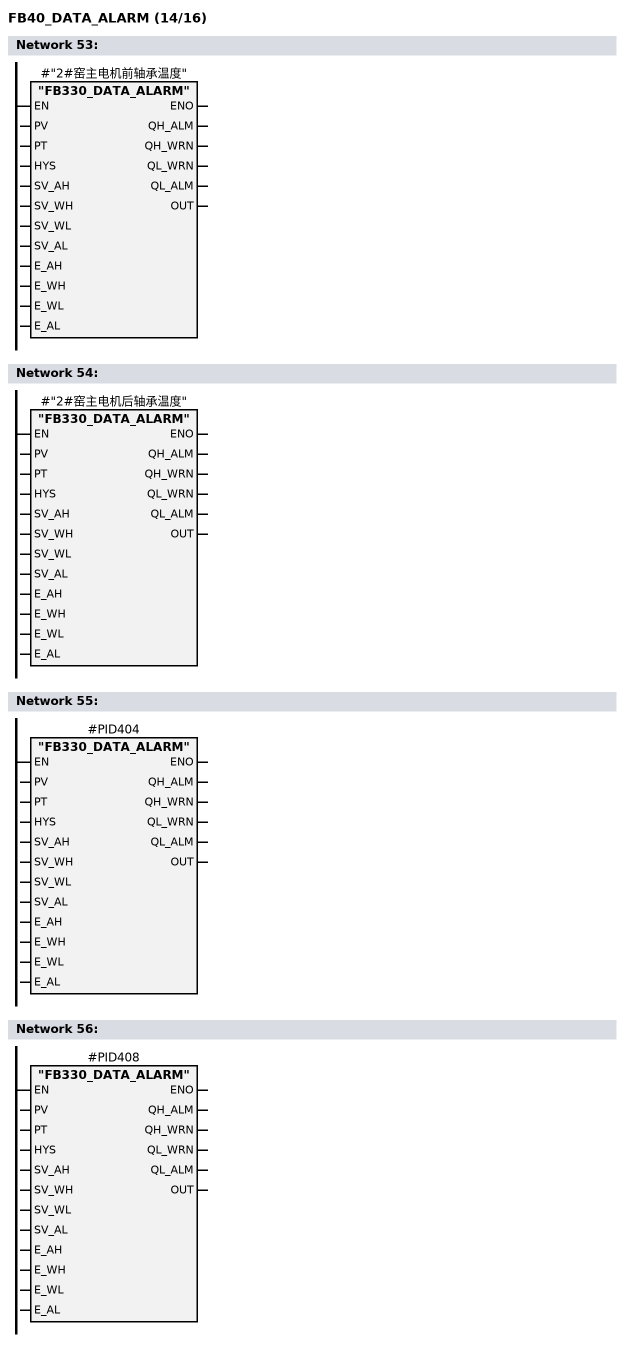
   RUNG wire#powerrail
      #"2#窑主电机前轴承温度"(PV :=, PT :=, HYS :=, SV_AH :=, SV_WH :=, SV_WL :=, SV_AL :=, E_AH :=, E_WH :=, E_WL :=, E_AL :=, QH_ALM =>, QH_WRN =>, QL_WRN =>, QL_ALM =>, OUT =>)
   END_RUNG
   // the same network as SCL:
   #"2#窑主电机前轴承温度"();   // "FB330_DATA_ALARM"
END_REGION

REGION Network 54
   RUNG wire#powerrail
      #"2#窑主电机后轴承温度"(PV :=, PT :=, HYS :=, SV_AH :=, SV_WH :=, SV_WL :=, SV_AL :=, E_AH :=, E_WH :=, E_WL :=, E_AL :=, QH_ALM =>, QH_WRN =>, QL_WRN =>, QL_ALM =>, OUT =>)
   END_RUNG
   // the same network as SCL:
   #"2#窑主电机后轴承温度"();   // "FB330_DATA_ALARM"
END_REGION

REGION Network 55
   RUNG wire#powerrail
      #PID404(PV :=, PT :=, HYS :=, SV_AH :=, SV_WH :=, SV_WL :=, SV_AL :=, E_AH :=, E_WH :=, E_WL :=, E_AL :=, QH_ALM =>, QH_WRN =>, QL_WRN =>, QL_ALM =>, OUT =>)
   END_RUNG
   // the same network as SCL:
   #PID404();   // "FB330_DATA_ALARM"
END_REGION

REGION Network 56
   RUNG wire#powerrail
      #PID408(PV :=, PT :=, HYS :=, SV_AH :=, SV_WH :=, SV_WL :=, SV_AL :=, E_AH :=, E_WH :=, E_WL :=, E_AL :=, QH_ALM =>, QH_WRN =>, QL_WRN =>, QL_ALM =>, OUT =>)
   END_RUNG
   // the same network as SCL:
   #PID408();   // "FB330_DATA_ALARM"
END_REGION

REGION Network 57
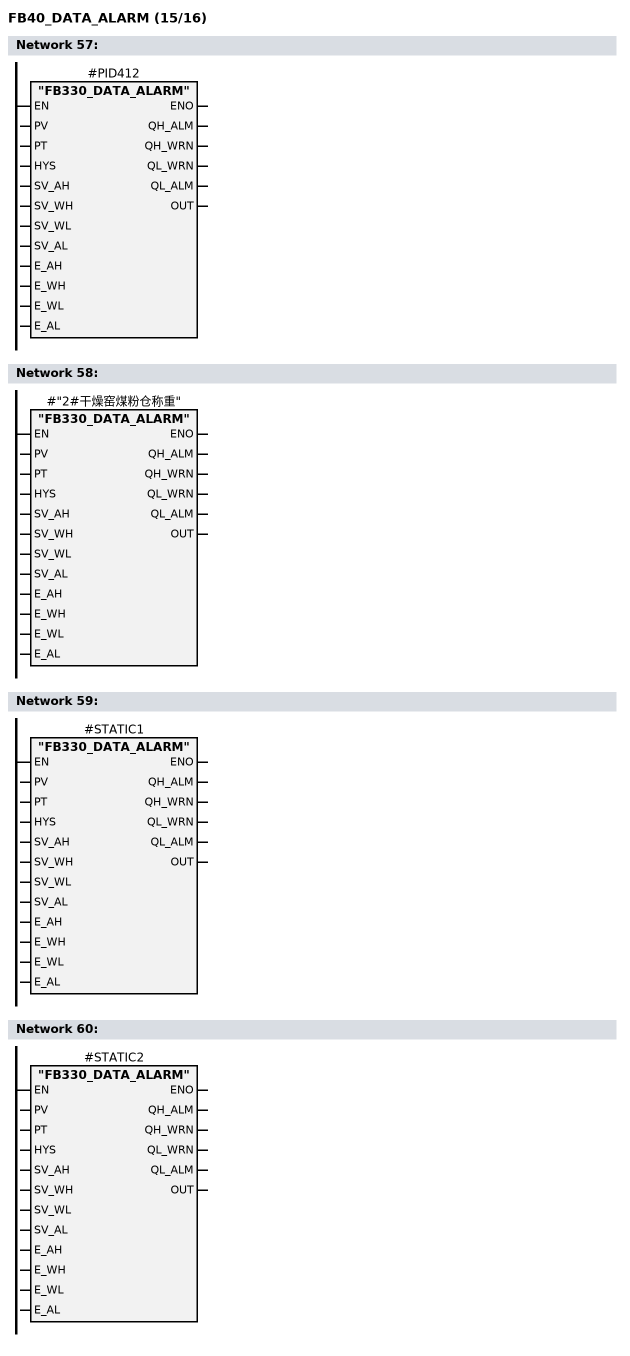
   RUNG wire#powerrail
      #PID412(PV :=, PT :=, HYS :=, SV_AH :=, SV_WH :=, SV_WL :=, SV_AL :=, E_AH :=, E_WH :=, E_WL :=, E_AL :=, QH_ALM =>, QH_WRN =>, QL_WRN =>, QL_ALM =>, OUT =>)
   END_RUNG
   // the same network as SCL:
   #PID412();   // "FB330_DATA_ALARM"
END_REGION

REGION Network 58
   RUNG wire#powerrail
      #"2#干燥窑煤粉仓称重"(PV :=, PT :=, HYS :=, SV_AH :=, SV_WH :=, SV_WL :=, SV_AL :=, E_AH :=, E_WH :=, E_WL :=, E_AL :=, QH_ALM =>, QH_WRN =>, QL_WRN =>, QL_ALM =>, OUT =>)
   END_RUNG
   // the same network as SCL:
   #"2#干燥窑煤粉仓称重"();   // "FB330_DATA_ALARM"
END_REGION

REGION Network 59
   RUNG wire#powerrail
      #STATIC1(PV :=, PT :=, HYS :=, SV_AH :=, SV_WH :=, SV_WL :=, SV_AL :=, E_AH :=, E_WH :=, E_WL :=, E_AL :=, QH_ALM =>, QH_WRN =>, QL_WRN =>, QL_ALM =>, OUT =>)
   END_RUNG
   // the same network as SCL:
   #STATIC1();   // "FB330_DATA_ALARM"
END_REGION

REGION Network 60
   RUNG wire#powerrail
      #STATIC2(PV :=, PT :=, HYS :=, SV_AH :=, SV_WH :=, SV_WL :=, SV_AL :=, E_AH :=, E_WH :=, E_WL :=, E_AL :=, QH_ALM =>, QH_WRN =>, QL_WRN =>, QL_ALM =>, OUT =>)
   END_RUNG
   // the same network as SCL:
   #STATIC2();   // "FB330_DATA_ALARM"
END_REGION

REGION Network 61
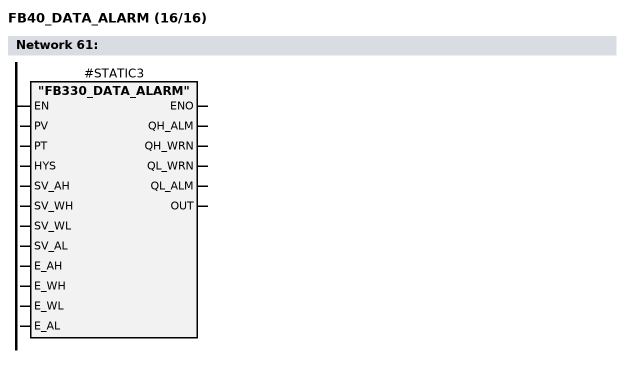
   RUNG wire#powerrail
      #STATIC3(PV :=, PT :=, HYS :=, SV_AH :=, SV_WH :=, SV_WL :=, SV_AL :=, E_AH :=, E_WH :=, E_WL :=, E_AL :=, QH_ALM =>, QH_WRN =>, QL_WRN =>, QL_ALM =>, OUT =>)
   END_RUNG
   // the same network as SCL:
   #STATIC3();   // "FB330_DATA_ALARM"
END_REGION
END_FUNCTION_BLOCK

FUNCTION_BLOCK "FB330_DATA_ALARM"   // FB330, LAD
{ S7_Optimized_Access := 'FALSE' }
VERSION : 0.1
// REAL的报警块
   VAR_INPUT
      PV : Real;   // 过程值
      PT : Real := 1.0;   // 系数
      HYS : Real;   // 回差值
      SV_AH : Real;   // 高报警设定值
      SV_WH : Real;   // 高警告设定值
      SV_WL : Real;   // 低警告设定值
      SV_AL : Real;   // 低报警设定值
      E_AH : Bool;   // 高报警使能
      E_WH : Bool;   // 高警告使能
      E_WL : Bool;   // 低警告使能
      E_AL : Bool;   // 低报警使能
   END_VAR
   VAR_OUTPUT
      QH_ALM : Bool;   // 高报警输出
      QH_WRN : Bool;   // 高警告输出
      QL_WRN : Bool;   // 低警告输出
      QL_ALM : Bool;   // 低报警输出
      OUT : Real;   // 输出
   END_VAR
   VAR
      SR1 : Bool;
      SR2 : Bool;
      SR3 : Bool;
      SR4 : Bool;
   END_VAR
   VAR_TEMP
      TEMP_AH : Real;
      TEMP_WH : Real;
      TEMP_AL : Real;
      TEMP_WL : Real;
      TEMP_OUT : Real;
   END_VAR
BEGIN

REGION Network 1
   // 系数转换
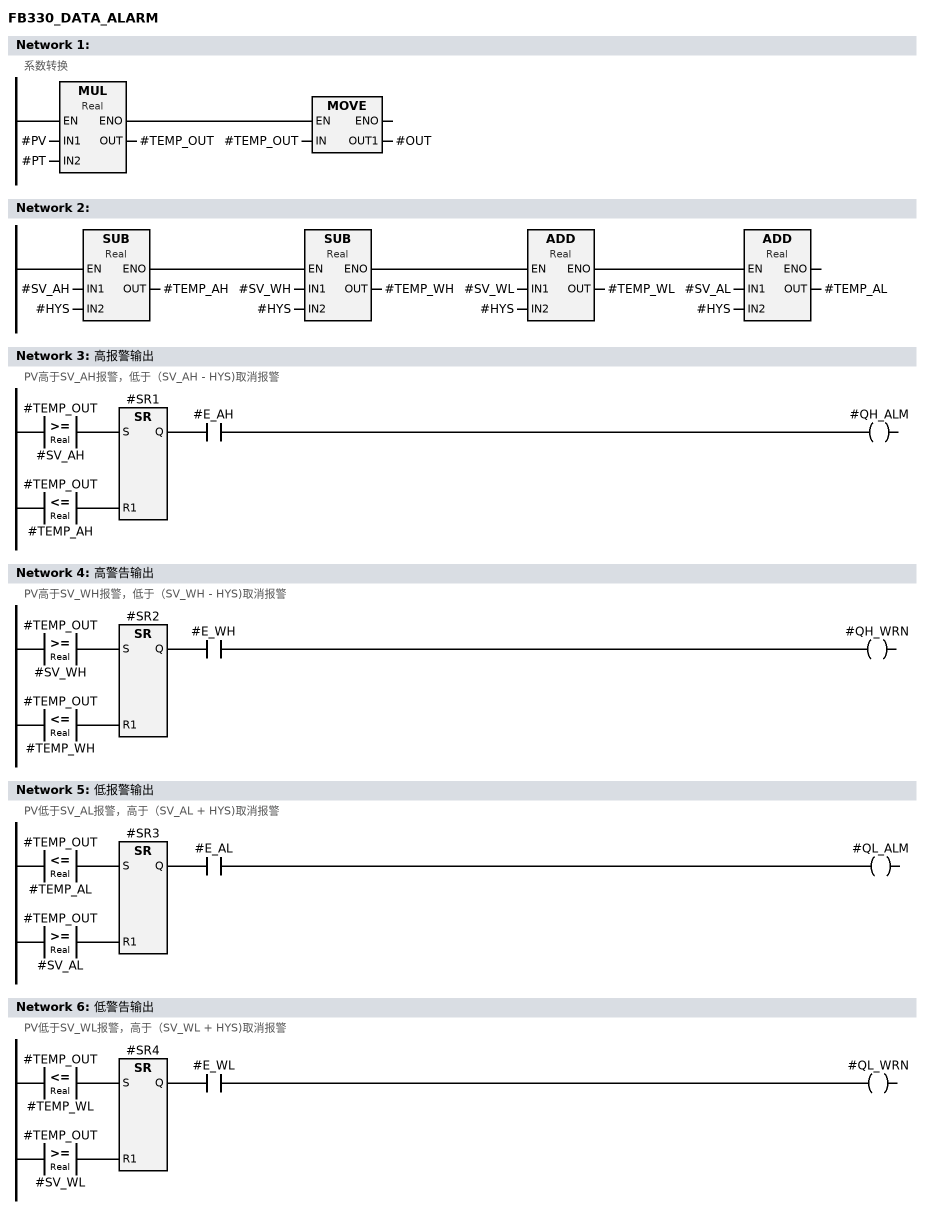
   RUNG wire#powerrail
      { S7_Templates := "SrcType := Real"; S7_GenerateENO := "TRUE" } Mul(in1 := #PV, in2 := #PT, out => #TEMP_OUT)
      { S7_GenerateENO := "TRUE" } Move(in := #TEMP_OUT, out1 => #OUT)
   END_RUNG
   // the same network as SCL:
   // ENO of a box is taken as its EN; it also drops when the box reports an error
   #TEMP_OUT := #PV * #PT;
   #OUT := #TEMP_OUT;
END_REGION

REGION Network 2
   RUNG wire#powerrail
      { S7_Templates := "SrcType := Real"; S7_GenerateENO := "TRUE" } Sub(in1 := #SV_AH, in2 := #HYS, out => #TEMP_AH)
      { S7_Templates := "SrcType := Real"; S7_GenerateENO := "TRUE" } Sub(in1 := #SV_WH, in2 := #HYS, out => #TEMP_WH)
      { S7_Templates := "SrcType := Real"; S7_GenerateENO := "TRUE" } Add(in1 := #SV_WL, in2 := #HYS, out => #TEMP_WL)
      { S7_Templates := "SrcType := Real"; S7_GenerateENO := "TRUE" } Add(in1 := #SV_AL, in2 := #HYS, out => #TEMP_AL)
   END_RUNG
   // the same network as SCL:
   // ENO of a box is taken as its EN; it also drops when the box reports an error
   #TEMP_AH := #SV_AH - #HYS;
   #TEMP_WH := #SV_WH - #HYS;
   #TEMP_WL := #SV_WL + #HYS;
   #TEMP_AL := #SV_AL + #HYS;
END_REGION

REGION Network 3: 高报警输出
   // PV高于SV_AH报警，低于（SV_AH - HYS)取消报警
   RUNG wire#powerrail
      { S7_Templates := "SrcType := Real" } GE_Contact(in1 := #TEMP_OUT, in2 := #SV_AH)
      S_SR(operand := #SR1, r1 := wire#w1)
      Contact( #E_AH )
      Coil( #QH_ALM )
   END_RUNG
   RUNG wire#powerrail
      { S7_Templates := "SrcType := Real" } LE_Contact(in1 := #TEMP_OUT, in2 := #TEMP_AH)
   END_RUNG wire#w1
   // the same network as SCL:
   IF #TEMP_OUT >= #SV_AH THEN
       #SR1 := TRUE;   // SR flip-flop
   END_IF;
   IF #TEMP_OUT <= #TEMP_AH THEN #SR1 := FALSE; END_IF;
   #QH_ALM := #SR1 AND #E_AH;
END_REGION

REGION Network 4: 高警告输出
   // PV高于SV_WH报警，低于（SV_WH - HYS)取消报警
   RUNG wire#powerrail
      { S7_Templates := "SrcType := Real" } GE_Contact(in1 := #TEMP_OUT, in2 := #SV_WH)
      S_SR(operand := #SR2, r1 := wire#w1)
      Contact( #E_WH )
      Coil( #QH_WRN )
   END_RUNG
   RUNG wire#powerrail
      { S7_Templates := "SrcType := Real" } LE_Contact(in1 := #TEMP_OUT, in2 := #TEMP_WH)
   END_RUNG wire#w1
   // the same network as SCL:
   IF #TEMP_OUT >= #SV_WH THEN
       #SR2 := TRUE;   // SR flip-flop
   END_IF;
   IF #TEMP_OUT <= #TEMP_WH THEN #SR2 := FALSE; END_IF;
   #QH_WRN := #SR2 AND #E_WH;
END_REGION

REGION Network 5: 低报警输出
   // PV低于SV_AL报警，高于（SV_AL + HYS)取消报警
   RUNG wire#powerrail
      { S7_Templates := "SrcType := Real" } LE_Contact(in1 := #TEMP_OUT, in2 := #TEMP_AL)
      S_SR(operand := #SR3, r1 := wire#w1)
      Contact( #E_AL )
      Coil( #QL_ALM )
   END_RUNG
   RUNG wire#powerrail
      { S7_Templates := "SrcType := Real" } GE_Contact(in1 := #TEMP_OUT, in2 := #SV_AL)
   END_RUNG wire#w1
   // the same network as SCL:
   IF #TEMP_OUT <= #TEMP_AL THEN
       #SR3 := TRUE;   // SR flip-flop
   END_IF;
   IF #TEMP_OUT >= #SV_AL THEN #SR3 := FALSE; END_IF;
   #QL_ALM := #SR3 AND #E_AL;
END_REGION

REGION Network 6: 低警告输出
   // PV低于SV_WL报警，高于（SV_WL + HYS)取消报警
   RUNG wire#powerrail
      { S7_Templates := "SrcType := Real" } LE_Contact(in1 := #TEMP_OUT, in2 := #TEMP_WL)
      S_SR(operand := #SR4, r1 := wire#w1)
      Contact( #E_WL )
      Coil( #QL_WRN )
   END_RUNG
   RUNG wire#powerrail
      { S7_Templates := "SrcType := Real" } GE_Contact(in1 := #TEMP_OUT, in2 := #SV_WL)
   END_RUNG wire#w1
   // the same network as SCL:
   IF #TEMP_OUT <= #TEMP_WL THEN
       #SR4 := TRUE;   // SR flip-flop
   END_IF;
   IF #TEMP_OUT >= #SV_WL THEN #SR4 := FALSE; END_IF;
   #QL_WRN := #SR4 AND #E_WL;
END_REGION
END_FUNCTION_BLOCK

FUNCTION_BLOCK "累计功能块2"   // FB333, LAD
{ S7_Optimized_Access := 'FALSE' }
VERSION : 0.1
   VAR_INPUT
      PV : Real;
      CLEAR1 : Bool;
      CLEAR2 : Bool;
      CLEAR3 : Bool;
      CLEAR4 : Bool;
   END_VAR
   VAR_OUTPUT
      OUT1 : Real;
      OUT2 : Real;
      OUT3 : Real;
      OUT4 : Real;
   END_VAR
   VAR
      "REAL" : Real;
      REAL1_1 : Real;
      REAL1_2 : Real;
      REAL1_3 : Real;
      REAL2_1 : Real;
      REAL2_2 : Real;
      REAL2_3 : Real;
      REAL3_1 : Real;
      REAL3_2 : Real;
      REAL3_3 : Real;
      REAL4_1 : Real;
      REAL4_2 : Real;
      REAL4_3 : Real;
      PV_DINT : DInt;
      DINT1 : DInt;
      DINT2 : DInt;
      DINT3 : DInt;
      DINT4 : DInt;
      P1 : Bool;
      P2 : Bool;
      P3 : Bool;
      P4 : Bool;
   END_VAR
   VAR_TEMP   // added for the SCL form of the ladder/FBD networks
      _w1 : Bool;
      _w2 : Bool;
   END_VAR
BEGIN

REGION Network 1
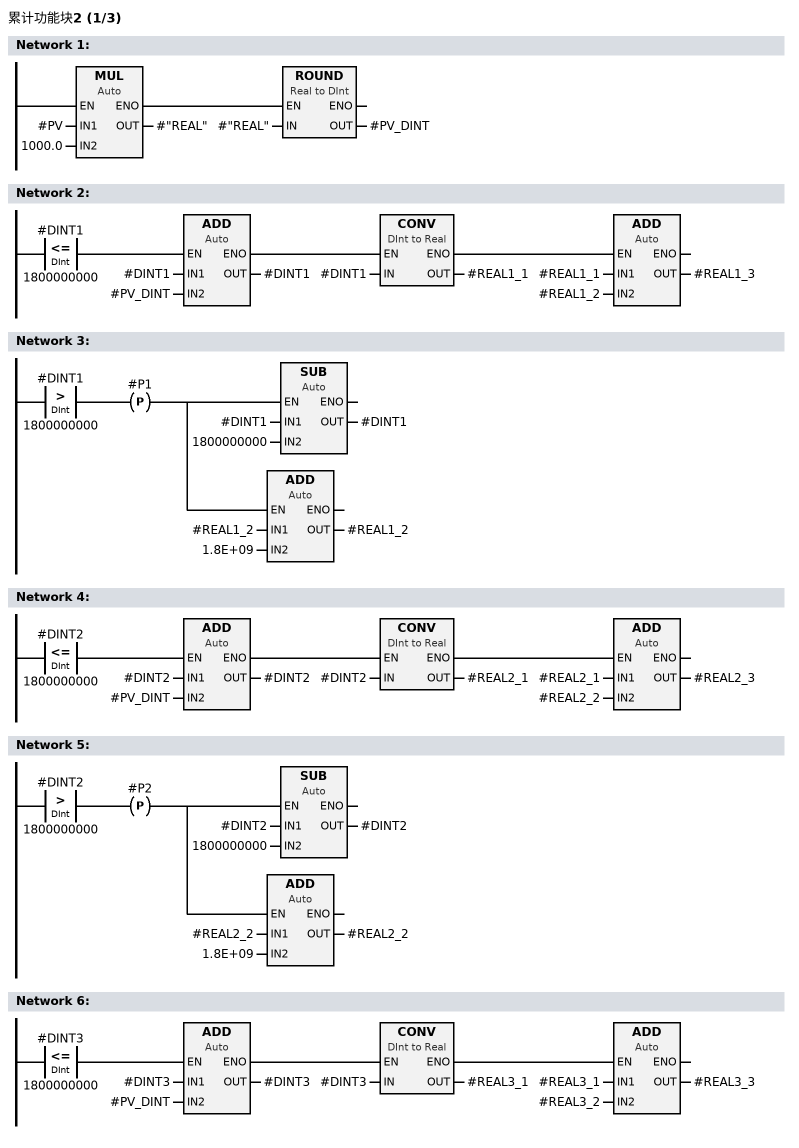
   RUNG wire#powerrail
      Mul(in1 := #PV, in2 := 1000.0, out => #"REAL")
      { S7_Templates := "[SrcType := Real, DestType := DInt]" } Round(in := #"REAL", out => #PV_DINT)
   END_RUNG
   // the same network as SCL:
   #"REAL" := #PV * 1000.0;
   #PV_DINT := ROUND(#"REAL");
END_REGION

REGION Network 2
   RUNG wire#powerrail
      { S7_Templates := "SrcType := DInt" } LE_Contact(in1 := #DINT1, in2 := 1800000000)
      Add(in1 := #DINT1, in2 := #PV_DINT, out => #DINT1)
      { S7_Templates := "[SrcType := DInt, DestType := Real]" } Convert(in := #DINT1, out => #REAL1_1)
      Add(in1 := #REAL1_1, in2 := #REAL1_2, out => #REAL1_3)
   END_RUNG
   // the same network as SCL:
   #_w1 := #DINT1 <= 1800000000;
   IF #_w1 THEN
       #DINT1 := #DINT1 + #PV_DINT;
       #REAL1_1 := DINT_TO_REAL(#DINT1);
       #REAL1_3 := #REAL1_1 + #REAL1_2;
   END_IF;
END_REGION

REGION Network 3
   RUNG wire#powerrail
      { S7_Templates := "SrcType := DInt" } GT_Contact(in1 := #DINT1, in2 := 1800000000)
      P_Trig( #P1 )
      wire#w1
      Sub(in1 := #DINT1, in2 := 1800000000, out => #DINT1)
   END_RUNG
   RUNG wire#w1
      Add(in1 := #REAL1_2, in2 := 1.8E+09, out => #REAL1_2)
   END_RUNG
   // the same network as SCL:
   #_w1 := #DINT1 > 1800000000;
   #_w2 := #_w1 AND NOT #P1;   // rising edge
   #P1 := #_w1;
   IF #_w2 THEN
       #DINT1 := #DINT1 - 1800000000;
       #REAL1_2 := #REAL1_2 + 1.8E+09;
   END_IF;
END_REGION

REGION Network 4
   RUNG wire#powerrail
      { S7_Templates := "SrcType := DInt" } LE_Contact(in1 := #DINT2, in2 := 1800000000)
      Add(in1 := #DINT2, in2 := #PV_DINT, out => #DINT2)
      { S7_Templates := "[SrcType := DInt, DestType := Real]" } Convert(in := #DINT2, out => #REAL2_1)
      Add(in1 := #REAL2_1, in2 := #REAL2_2, out => #REAL2_3)
   END_RUNG
   // the same network as SCL:
   #_w1 := #DINT2 <= 1800000000;
   IF #_w1 THEN
       #DINT2 := #DINT2 + #PV_DINT;
       #REAL2_1 := DINT_TO_REAL(#DINT2);
       #REAL2_3 := #REAL2_1 + #REAL2_2;
   END_IF;
END_REGION

REGION Network 5
   RUNG wire#powerrail
      { S7_Templates := "SrcType := DInt" } GT_Contact(in1 := #DINT2, in2 := 1800000000)
      P_Trig( #P2 )
      wire#w1
      Sub(in1 := #DINT2, in2 := 1800000000, out => #DINT2)
   END_RUNG
   RUNG wire#w1
      Add(in1 := #REAL2_2, in2 := 1.8E+09, out => #REAL2_2)
   END_RUNG
   // the same network as SCL:
   #_w1 := #DINT2 > 1800000000;
   #_w2 := #_w1 AND NOT #P2;   // rising edge
   #P2 := #_w1;
   IF #_w2 THEN
       #DINT2 := #DINT2 - 1800000000;
       #REAL2_2 := #REAL2_2 + 1.8E+09;
   END_IF;
END_REGION

REGION Network 6
   RUNG wire#powerrail
      { S7_Templates := "SrcType := DInt" } LE_Contact(in1 := #DINT3, in2 := 1800000000)
      Add(in1 := #DINT3, in2 := #PV_DINT, out => #DINT3)
      { S7_Templates := "[SrcType := DInt, DestType := Real]" } Convert(in := #DINT3, out => #REAL3_1)
      Add(in1 := #REAL3_1, in2 := #REAL3_2, out => #REAL3_3)
   END_RUNG
   // the same network as SCL:
   #_w1 := #DINT3 <= 1800000000;
   IF #_w1 THEN
       #DINT3 := #DINT3 + #PV_DINT;
       #REAL3_1 := DINT_TO_REAL(#DINT3);
       #REAL3_3 := #REAL3_1 + #REAL3_2;
   END_IF;
END_REGION

REGION Network 7
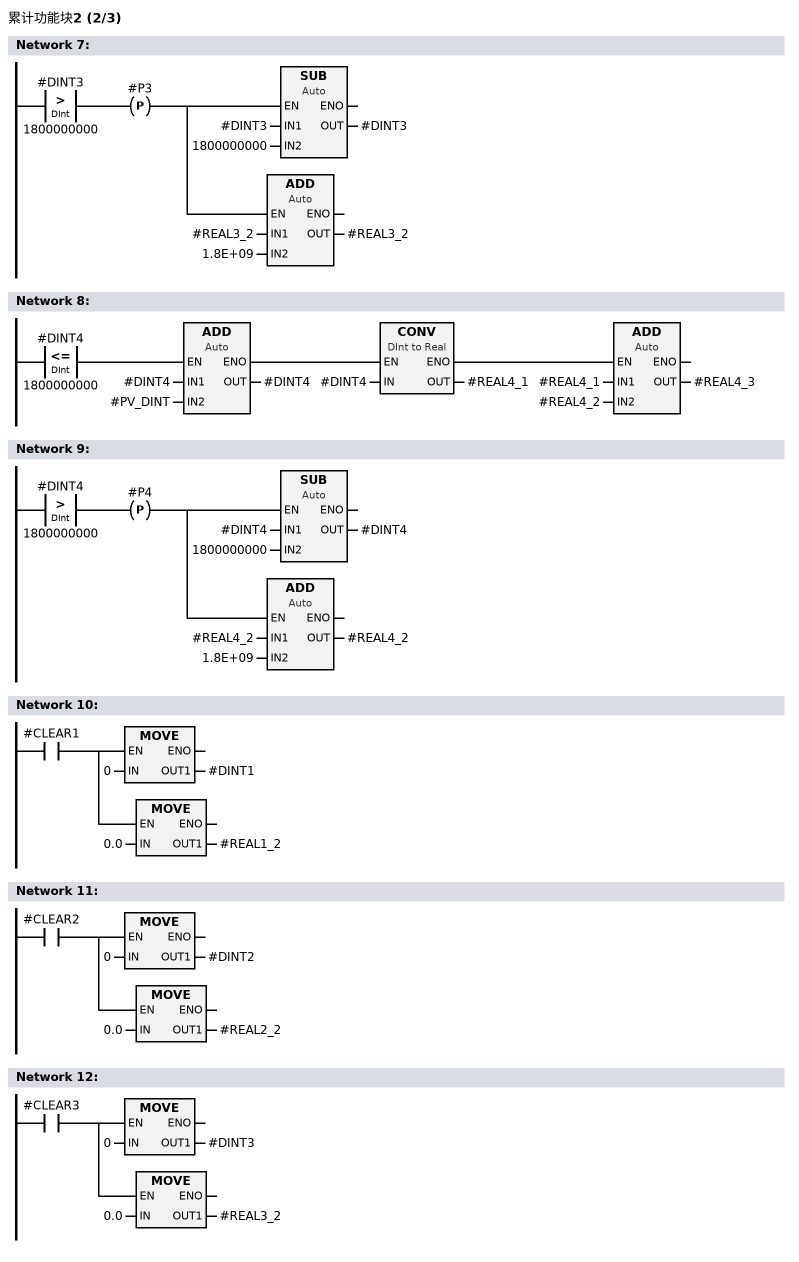
   RUNG wire#powerrail
      { S7_Templates := "SrcType := DInt" } GT_Contact(in1 := #DINT3, in2 := 1800000000)
      P_Trig( #P3 )
      wire#w1
      Sub(in1 := #DINT3, in2 := 1800000000, out => #DINT3)
   END_RUNG
   RUNG wire#w1
      Add(in1 := #REAL3_2, in2 := 1.8E+09, out => #REAL3_2)
   END_RUNG
   // the same network as SCL:
   #_w1 := #DINT3 > 1800000000;
   #_w2 := #_w1 AND NOT #P3;   // rising edge
   #P3 := #_w1;
   IF #_w2 THEN
       #DINT3 := #DINT3 - 1800000000;
       #REAL3_2 := #REAL3_2 + 1.8E+09;
   END_IF;
END_REGION

REGION Network 8
   RUNG wire#powerrail
      { S7_Templates := "SrcType := DInt" } LE_Contact(in1 := #DINT4, in2 := 1800000000)
      Add(in1 := #DINT4, in2 := #PV_DINT, out => #DINT4)
      { S7_Templates := "[SrcType := DInt, DestType := Real]" } Convert(in := #DINT4, out => #REAL4_1)
      Add(in1 := #REAL4_1, in2 := #REAL4_2, out => #REAL4_3)
   END_RUNG
   // the same network as SCL:
   #_w1 := #DINT4 <= 1800000000;
   IF #_w1 THEN
       #DINT4 := #DINT4 + #PV_DINT;
       #REAL4_1 := DINT_TO_REAL(#DINT4);
       #REAL4_3 := #REAL4_1 + #REAL4_2;
   END_IF;
END_REGION

REGION Network 9
   RUNG wire#powerrail
      { S7_Templates := "SrcType := DInt" } GT_Contact(in1 := #DINT4, in2 := 1800000000)
      P_Trig( #P4 )
      wire#w1
      Sub(in1 := #DINT4, in2 := 1800000000, out => #DINT4)
   END_RUNG
   RUNG wire#w1
      Add(in1 := #REAL4_2, in2 := 1.8E+09, out => #REAL4_2)
   END_RUNG
   // the same network as SCL:
   #_w1 := #DINT4 > 1800000000;
   #_w2 := #_w1 AND NOT #P4;   // rising edge
   #P4 := #_w1;
   IF #_w2 THEN
       #DINT4 := #DINT4 - 1800000000;
       #REAL4_2 := #REAL4_2 + 1.8E+09;
   END_IF;
END_REGION

REGION Network 10
   RUNG wire#powerrail
      Contact( #CLEAR1 )
      wire#w1
      Move(in := 0, out1 => #DINT1)
   END_RUNG
   RUNG wire#w1
      Move(in := 0.0, out1 => #REAL1_2)
   END_RUNG
   // the same network as SCL:
   IF #CLEAR1 THEN
       #DINT1 := 0;
       #REAL1_2 := 0.0;
   END_IF;
END_REGION

REGION Network 11
   RUNG wire#powerrail
      Contact( #CLEAR2 )
      wire#w1
      Move(in := 0, out1 => #DINT2)
   END_RUNG
   RUNG wire#w1
      Move(in := 0.0, out1 => #REAL2_2)
   END_RUNG
   // the same network as SCL:
   IF #CLEAR2 THEN
       #DINT2 := 0;
       #REAL2_2 := 0.0;
   END_IF;
END_REGION

REGION Network 12
   RUNG wire#powerrail
      Contact( #CLEAR3 )
      wire#w1
      Move(in := 0, out1 => #DINT3)
   END_RUNG
   RUNG wire#w1
      Move(in := 0.0, out1 => #REAL3_2)
   END_RUNG
   // the same network as SCL:
   IF #CLEAR3 THEN
       #DINT3 := 0;
       #REAL3_2 := 0.0;
   END_IF;
END_REGION

REGION Network 13
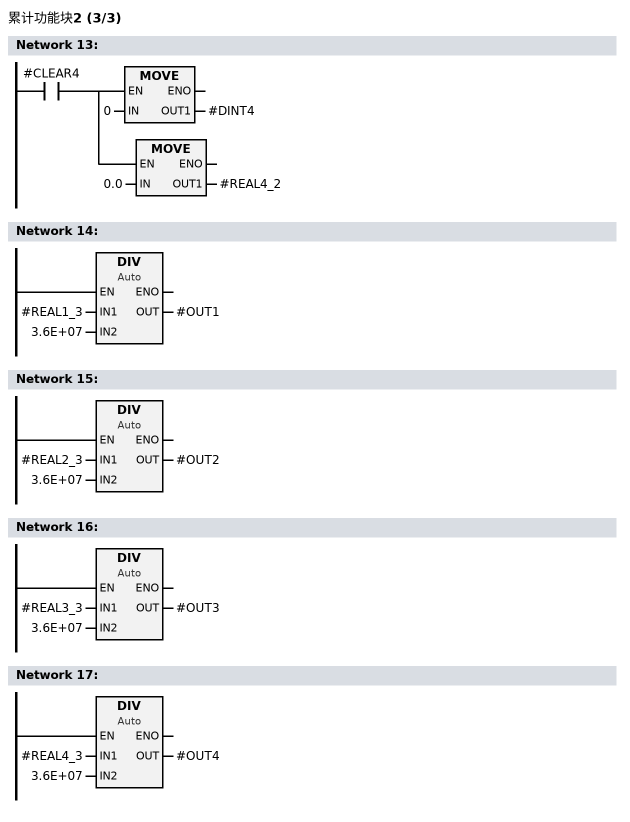
   RUNG wire#powerrail
      Contact( #CLEAR4 )
      wire#w1
      Move(in := 0, out1 => #DINT4)
   END_RUNG
   RUNG wire#w1
      Move(in := 0.0, out1 => #REAL4_2)
   END_RUNG
   // the same network as SCL:
   IF #CLEAR4 THEN
       #DINT4 := 0;
       #REAL4_2 := 0.0;
   END_IF;
END_REGION

REGION Network 14
   RUNG wire#powerrail
      Div(in1 := #REAL1_3, in2 := 3.6E+07, out => #OUT1)
   END_RUNG
   // the same network as SCL:
   #OUT1 := #REAL1_3 / 3.6E+07;
END_REGION

REGION Network 15
   RUNG wire#powerrail
      Div(in1 := #REAL2_3, in2 := 3.6E+07, out => #OUT2)
   END_RUNG
   // the same network as SCL:
   #OUT2 := #REAL2_3 / 3.6E+07;
END_REGION

REGION Network 16
   RUNG wire#powerrail
      Div(in1 := #REAL3_3, in2 := 3.6E+07, out => #OUT3)
   END_RUNG
   // the same network as SCL:
   #OUT3 := #REAL3_3 / 3.6E+07;
END_REGION

REGION Network 17
   RUNG wire#powerrail
      Div(in1 := #REAL4_3, in2 := 3.6E+07, out => #OUT4)
   END_RUNG
   // the same network as SCL:
   #OUT4 := #REAL4_3 / 3.6E+07;
END_REGION
END_FUNCTION_BLOCK

FUNCTION "电机块" : Void   // FC1, LAD
{ S7_Optimized_Access := 'FALSE' }
VERSION : 0.1
   VAR_INPUT
      ST : Bool;
      LR : Bool;
      STP : Bool;
      FAULT : Bool;
   END_VAR
   VAR_IN_OUT
      OUT : Bool;
   END_VAR
BEGIN

REGION Network 1
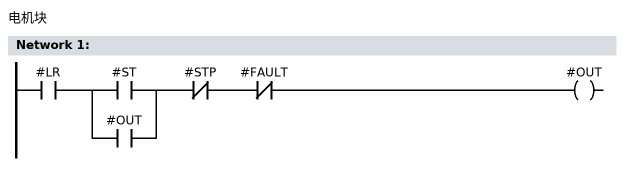
   RUNG wire#powerrail
      Contact( #LR )
      wire#w1
      Contact( #ST )
      wire#w2
      I_Contact( #STP )
      I_Contact( #FAULT )
      Coil( #OUT )
   END_RUNG
   RUNG wire#w1
      Contact( #OUT )
   END_RUNG wire#w2
   // the same network as SCL:
   #OUT := #LR AND (#ST OR #OUT) AND NOT #STP AND NOT #FAULT;
END_REGION
END_FUNCTION

FUNCTION "风机" : Void   // FC2, LAD
{ S7_Optimized_Access := 'FALSE' }
VERSION : 0.1
BEGIN

REGION Network 1
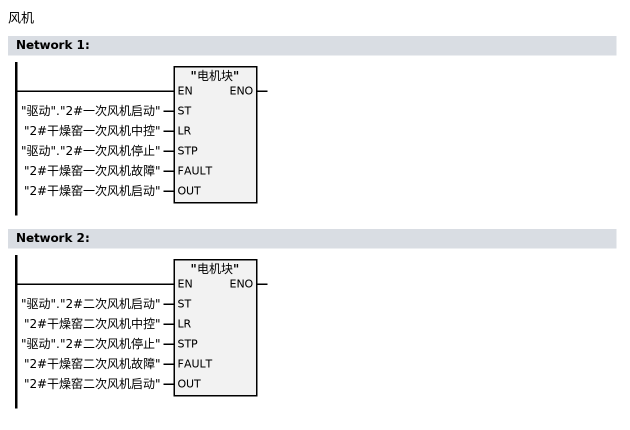
   RUNG wire#powerrail
      "电机块"(ST := "驱动"."2#一次风机启动", LR := "2#干燥窑一次风机中控", STP := "驱动"."2#一次风机停止", FAULT := "2#干燥窑一次风机故障", OUT := "2#干燥窑一次风机启动")
   END_RUNG
   // the same network as SCL:
   "电机块"(ST := "驱动"."2#一次风机启动",
         LR := "2#干燥窑一次风机中控",
         STP := "驱动"."2#一次风机停止",
         FAULT := "2#干燥窑一次风机故障",
         OUT := "2#干燥窑一次风机启动");
END_REGION

REGION Network 2
   RUNG wire#powerrail
      "电机块"(ST := "驱动"."2#二次风机启动", LR := "2#干燥窑二次风机中控", STP := "驱动"."2#二次风机停止", FAULT := "2#干燥窑二次风机故障", OUT := "2#干燥窑二次风机启动")
   END_RUNG
   // the same network as SCL:
   "电机块"(ST := "驱动"."2#二次风机启动",
         LR := "2#干燥窑二次风机中控",
         STP := "驱动"."2#二次风机停止",
         FAULT := "2#干燥窑二次风机故障",
         OUT := "2#干燥窑二次风机启动");
END_REGION
END_FUNCTION

FUNCTION "程序" : Void   // FC3, LAD
{ S7_Optimized_Access := 'FALSE' }
VERSION : 0.1
   VAR_TEMP   // added for the SCL form of the ladder/FBD networks
      _w1 : Bool;
      _s5time1 : S5Time;
   END_VAR
BEGIN

REGION Network 1
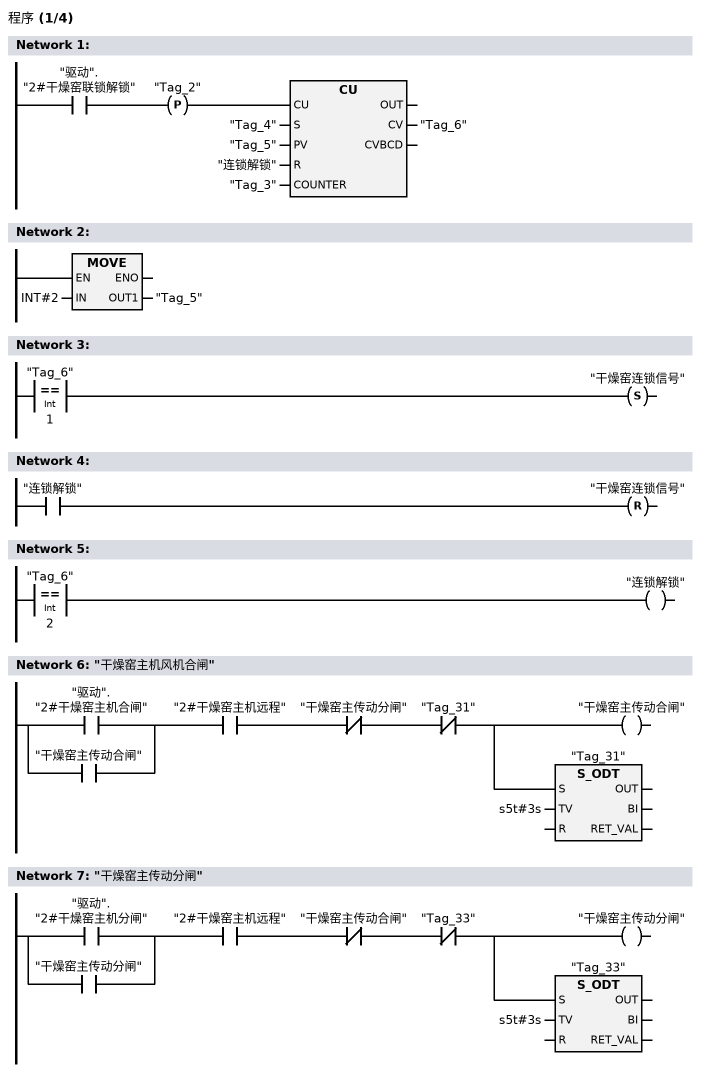
   // no SCL statement known for Cu: written as a call
   #_w1 := "驱动"."2#干燥窑联锁解锁" AND NOT "Tag_2";   // rising edge
   "Tag_2" := "驱动"."2#干燥窑联锁解锁";
   Cu(cu := #_w1, s := "Tag_4", pv := "Tag_5", r := "连锁解锁", "counter" := "Tag_3", cv => "Tag_6");
END_REGION

REGION Network 2
   RUNG wire#powerrail
      { S7_GenerateENO := "TRUE" } Move(in := INT#2, out1 => "Tag_5")
   END_RUNG
   // the same network as SCL:
   "Tag_5" := INT#2;
END_REGION

REGION Network 3
   RUNG wire#powerrail
      { S7_Templates := "SrcType := Int" } EQ_Contact(in1 := "Tag_6", in2 := 1)
      S_Coil( "干燥窑连锁信号" )
   END_RUNG
   // the same network as SCL:
   IF "Tag_6" = 1 THEN "干燥窑连锁信号" := TRUE; END_IF;
END_REGION

REGION Network 4
   RUNG wire#powerrail
      Contact( "连锁解锁" )
      R_Coil( "干燥窑连锁信号" )
   END_RUNG
   // the same network as SCL:
   IF "连锁解锁" THEN "干燥窑连锁信号" := FALSE; END_IF;
END_REGION

REGION Network 5
   RUNG wire#powerrail
      { S7_Templates := "SrcType := Int" } EQ_Contact(in1 := "Tag_6", in2 := 2)
      Coil( "连锁解锁" )
   END_RUNG
   // the same network as SCL:
   "连锁解锁" := "Tag_6" = 2;
END_REGION

REGION Network 6: "干燥窑主机风机合闸"
   RUNG wire#powerrail
      Contact( "驱动"."2#干燥窑主机合闸" )
      wire#w1
      Contact( "2#干燥窑主机远程" )
      I_Contact( "干燥窑主传动分闸" )
      I_Contact( "Tag_31" )
      wire#w2
      Coil( "干燥窑主传动合闸" )
   END_RUNG
   RUNG wire#powerrail
      Contact( "干燥窑主传动合闸" )
   END_RUNG wire#w1
   RUNG wire#w2
      S_ODT(T_NO := "Tag_31", TV := s5t#3s, R :=, BI =>, RET_VAL =>)
   END_RUNG
   // the same network as SCL:
   "干燥窑主传动合闸" := ("驱动"."2#干燥窑主机合闸" OR "干燥窑主传动合闸") AND "2#干燥窑主机远程" AND NOT "干燥窑主传动分闸" AND NOT "Tag_31";
   #_s5time1 := S_ODT(T_NO := "Tag_31", S := "干燥窑主传动合闸", TV := s5t#3s);
END_REGION

REGION Network 7: "干燥窑主传动分闸"
   RUNG wire#powerrail
      Contact( "驱动"."2#干燥窑主机分闸" )
      wire#w1
      Contact( "2#干燥窑主机远程" )
      I_Contact( "干燥窑主传动合闸" )
      I_Contact( "Tag_33" )
      wire#w2
      Coil( "干燥窑主传动分闸" )
   END_RUNG
   RUNG wire#powerrail
      Contact( "干燥窑主传动分闸" )
   END_RUNG wire#w1
   RUNG wire#w2
      S_ODT(T_NO := "Tag_33", TV := s5t#3s, R :=, BI =>, RET_VAL =>)
   END_RUNG
   // the same network as SCL:
   "干燥窑主传动分闸" := ("驱动"."2#干燥窑主机分闸" OR "干燥窑主传动分闸") AND "2#干燥窑主机远程" AND NOT "干燥窑主传动合闸" AND NOT "Tag_33";
   #_s5time1 := S_ODT(T_NO := "Tag_33", S := "干燥窑主传动分闸", TV := s5t#3s);
END_REGION

REGION Network 8
